
               #State_DwellAndReOx_SupplyToDeck:
                   IF #DECK_MANAGE_START_SUPPLY.ShutdownDemand THEN
                       #State.System := #State_Shutdown;
                   ELSIF "1092_HMI_OP_FLAGS".DeckSupplyOk THEN
                       #State.ReOx := #State_DwellAndReOx_OpenPVV;
                   ELSE
                       #DECK_MANAGE_START_SUPPLY();
                       "58_INTRNL_COMMS".BWT_TO_GCU.SPLY_GAS := True;
                       "58_INTRNL_COMMS".BWT_TO_GCU.STP_GAS := False;
                   END_IF;
               #State_DwellAndReOx_OpenPVV:
                   IF "1090_HMI_IP_FLAGS".PressVacuumValves THEN
                       #State.ReOx := #State_DwellAndReOx_OpenGTT;
                   ELSE
                       #NextStageCheck := "1151_NEXT_STAGE_CHECK_PVV"(AlarmState := #State_Shutdown, PVVX_OUT := #PVVX_OUT, State := #State, TankData := #TankData);
                       IF #NextStageCheck.Demand_Complete AND NOT #NextStageCheck.Alarm_Active THEN
                           #State.ReOx := #State_DwellAndReOx_OpenGTT;
                       END_IF;
                   END_IF;
               #State_DwellAndReOx_OpenGTT:
                   #NextStageCheck := "1150_NEXT_STAGE_CHECK_GTT"(AlarmState := #State_Shutdown, GTT_OUT := #GTT_OUT, State := #State, TankData := #TankData);
                   IF #NextStageCheck.Demand_Complete AND NOT #NextStageCheck.Alarm_Active THEN
                       #State.ReOx := #State_DwellAndReOx_Monitor;
                       "1134_MOVE_TANKS_INGROUP_NEW_STATE"(TankData := #TankData,
                                                          State := #State,
                                                          NewState := #TankState_ReOx);
                       // Reset timer information for this new treatment group
                       #XEOX_TIMER(IN := False,
                                   PT := "1190_FIXED_CONSTANTS".ReOxMin_Time,
                                   R := True);
                       #XEOX_PAUSE_TIMER(IN := False,
                                         PT := #MaxTimerPT,
                                         R := True);
                       #XEOX_PausedTime := LT#0s;
                   END_IF;
               #State_DwellAndReOx_Monitor:
                   IF #XEOX_TIMER.Q THEN
                       #NextStageCheck := "1153_NEXT_STAGE_CHECK_XEOX"(AlarmState := #State_Shutdown, State := #State, TankData := #TankData);
                       IF #NextStageCheck.Demand_Complete AND NOT #NextStageCheck.Alarm_Active THEN
                           #NextTreatmentGroup := "1136_CALC_NEXT_TREATMENT_GROUP"(NumberOfTreatmentGroups := "1190_FIXED_CONSTANTS".NumberOfTreatmentGroups, State := #State, TankData := #TankData);
                           IF #NextTreatmentGroup = -1 THEN
                               #DECK_MANAGE_STOP_SUPPLY.Stage := 0;
                               #State.ReOx := #State_DwellAndReOx_StopSupplyToDeck;
                           ELSE
                               #State.ReOx := #State_DwellAndReOx_CloseGTT;
                           END_IF;
                       END_IF;
                   ELSE
                       IF "58_INTRNL_COMMS".GCU_TO_BWT.GAS_AVLBL THEN
                           // continue counting on the reox timer as GCU is in a healthy state.
                           // increment the paused time as this shall be added to the deoxmin_time due to stoppage.
                           #XEOX_PausedTime += #XEOX_PAUSE_TIMER.ET;
                           #XEOX_TIMER(IN := True,
                                       PT := "1190_FIXED_CONSTANTS".ReOxMin_Time + #XEOX_PausedTime,
                                       R := False);
                           // keep XEOX pause timer in reset state.
                           #XEOX_PAUSE_TIMER(IN := False,
                                             PT := #MaxTimerPT,
                                             R := True);
                       ELSE
                           // Keep reox timer paused, whilst pause timer increments.
                           #XEOX_TIMER(IN := False,
                                       PT := "1190_FIXED_CONSTANTS".ReOxMin_Time + #XEOX_PausedTime,
                                       R := False);
                           #XEOX_PAUSE_TIMER(IN := True,
                                             PT := #MaxTimerPT,
                                             R := False);
                       END_IF;
                   END_IF;
               #State_DwellAndReOx_CloseGTT:
                   #NextStageCheck := "1150_NEXT_STAGE_CHECK_GTT"(AlarmState := #State_Shutdown, GTT_OUT := #GTT_OUT, State := #State, TankData := #TankData);
                   IF #NextStageCheck.Demand_Complete AND NOT #NextStageCheck.Alarm_Active THEN
                       // All tanks in this treatment group are now re-oxed, move them to post-dwell tank state.
                       "1134_MOVE_TANKS_INGROUP_NEW_STATE"(TankData := #TankData,
                                                          State := #State,
                                                          NewState := #TankState_PostDwell);
                      #NextTreatmentGroup := "1136_CALC_NEXT_TREATMENT_GROUP"(NumberOfTreatmentGroups := "1190_FIXED_CONSTANTS".NumberOfTreatmentGroups, State := #State, TankData := #TankData);
                       IF #NextTreatmentGroup = -1 THEN
                           #State.TreatmentGroup := 1;
                           #State.System := #State_DwellAndComplete;
                           #State.Complete := #State_DwellAndComplete_WaitPostDwell;
                       ELSE
                           // Are there more treatment groups to go? If so, restart the ReOx process on the next treatment group.
                           #State.TreatmentGroup := #NextTreatmentGroup;
                           #State.ReOx := #State_DwellAndReOx_WaitMidDwell;
                       END_IF;
                   END_IF;
               #State_DwellAndReOx_StopSupplyToDeck:
                   IF #DECK_MANAGE_STOP_SUPPLY.ShutdownDemand THEN
                       // Deck supply has failed, shutdown demand.
                       #State.System := #State_Shutdown;
                   ELSIF #DECK_MANAGE_STOP_SUPPLY.StopDeckSupplyDone THEN
                       // Deck stop supply is complete, go back to close the final set of GTT valves.
                       #State.ReOx := #State_DwellAndReOx_CloseGTT;
                   ELSE
                       // Deck stop supply is not complete yet, run stop supply to deck automation.
                       #DECK_MANAGE_STOP_SUPPLY();
                       "58_INTRNL_COMMS".BWT_TO_GCU.SPLY_GAS := False;
                       "58_INTRNL_COMMS".BWT_TO_GCU.STP_GAS := True;
                   END_IF;
           END_CASE;

       #State_DwellAndComplete:
           CASE #State.Complete OF
               #State_DwellAndComplete_WaitPostDwell:
                   #NextStageCheck := "1152_NEXT_STAGE_CHECK_TIMER"(AlarmState := #State_Shutdown, State := #State, TankData := #TankData);
                   IF #NextStageCheck.Demand_Complete AND NOT #NextStageCheck.Alarm_Active THEN
                       "1134_MOVE_TANKS_INGROUP_NEW_STATE"(TankData := #TankData,
                                                          State := #State,
                                                          NewState := #TankState_Done);
                      #NextTreatmentGroup := "1136_CALC_NEXT_TREATMENT_GROUP"(NumberOfTreatmentGroups := "1190_FIXED_CONSTANTS".NumberOfTreatmentGroups, State := #State, TankData := #TankData);
                       IF #NextTreatmentGroup = -1 THEN
                           #State.Complete := #State_DwellAndComplete_Done;
                       ELSE
                           // Are there more treatment groups to go? If so, wait for the next treatment group to finish post-dwell.
                           #State.TreatmentGroup := #NextTreatmentGroup;
                           #State.Complete := #State_DwellAndComplete_WaitPostDwell;
                       END_IF;
                   END_IF;
               #State_DwellAndComplete_Done:
                   // At this stage, all tanks have been processed.
                   "1092_HMI_OP_FLAGS".HMI_Warnings.Active := True;
                   "1092_HMI_OP_FLAGS".HMI_Warnings.Message := 'Ballast Water Treatment process has completed. All active tanks have been treated.';
           END_CASE;
       #State_Shutdown:
           "58_INTRNL_COMMS".BWT_TO_GCU.SHT_DN := True;
           IF #ShutdownStageReset THEN
               // If this is the first call to the shutdown, reset the stage to zero
               // do not call this reset again once called once.
               #DECK_MANAGE_STOP_SUPPLY.Stage := 0;
               #ShutdownStageReset := false;
           END_IF;
           IF #DECK_MANAGE_STOP_SUPPLY.ShutdownDemand THEN
               // Deck supply has failed, shutdown demand.6000
               #State.System := #State_Shutdown;
               "1092_HMI_OP_FLAGS".HMI_Warnings.Active := True;
               "1092_HMI_OP_FLAGS".HMI_Warnings.Message := 'BWTS Shutdown: failed to stop supply to main deck';
           ELSIF #DECK_MANAGE_STOP_SUPPLY.StopDeckSupplyDone THEN
               "1092_HMI_OP_FLAGS".HMI_Warnings.Active := True;
               "1092_HMI_OP_FLAGS".HMI_Warnings.Message := 'BWTS Shutdown: maain deck supply stopped';
           ELSE
               // Deck stop supply is not complete yet, run stop supply to deck automation.
               "1092_HMI_OP_FLAGS".HMI_Warnings.Active := True;
               "1092_HMI_OP_FLAGS".HMI_Warnings.Message := 'BWTS Shutdown: closing main line to deck';
               #DECK_MANAGE_STOP_SUPPLY();
           END_IF;
   END_CASE;

   (*
       Set all actuate commands to false to initialise on each scan cycle. Therefore each tank must now
       confirm that it wants the valve in question to actuate. Then call each tank in turn, make control
       decisions based on 1. The tank sub-state, the system operating state (and subsequently, deox/reox
       states if applicable.
   *)
   FOR #Index := 1 TO #NumberOfTanks DO
       #GTT_IN.GTT_Actuate[#Index] := False;
       #PVVX_IN.PVVx_Actuate[#Index] := False;
   END_FOR;
   #TANK_CONTROL_FPT(State := #State,
                     PVVX_IN := #PVVX_IN,
                     GTT_IN := #GTT_IN,
                     PVVX_OUT_DATA := #PVVX_OUT,
                     GTT_OUT_DATA := #GTT_OUT,
                     TankData := #TankData[1],
                     TankIPData := "20_TANKS_IP_DATA".RIO_01.FIRST_TANK);
   #TANK_CONTROL_1P(State := #State,
                    PVVX_IN := #PVVX_IN,
                    GTT_IN := #GTT_IN,
                    PVVX_OUT_DATA := #PVVX_OUT,
                    GTT_OUT_DATA := #GTT_OUT,
                    TankData := #TankData[2],
                    TankIPData := "20_TANKS_IP_DATA".RIO_01.SECOND_TANK);
   #TANK_CONTROL_1S(State := #State,
                    PVVX_IN := #PVVX_IN,
                    GTT_IN := #GTT_IN,
                    PVVX_OUT_DATA := #PVVX_OUT,
                    GTT_OUT_DATA := #GTT_OUT,
                    TankData := #TankData[3],
                    TankIPData := "20_TANKS_IP_DATA".RIO_01.THIRD_TANK);
   #TANK_CONTROL_2P(State := #State,
                    PVVX_IN := #PVVX_IN,
                    GTT_IN := #GTT_IN,
                    PVVX_OUT_DATA := #PVVX_OUT,
                    GTT_OUT_DATA := #GTT_OUT,
                    TankData := #TankData[4],
                    TankIPData := "20_TANKS_IP_DATA".RIO_02.FIRST_TANK);
   #TANK_CONTROL_2S(State := #State,
                    PVVX_IN := #PVVX_IN,
                    GTT_IN := #GTT_IN,
                    PVVX_OUT_DATA := #PVVX_OUT,
                    GTT_OUT_DATA := #GTT_OUT,
                    TankData := #TankData[5],
                    TankIPData := "20_TANKS_IP_DATA".RIO_02.SECOND_TANK);
   #TANK_CONTROL_3P(State := #State,
                    PVVX_IN := #PVVX_IN,
                    GTT_IN := #GTT_IN,
                    PVVX_OUT_DATA := #PVVX_OUT,
                    GTT_OUT_DATA := #GTT_OUT,
                    TankData := #TankData[6],
                    TankIPData := "20_TANKS_IP_DATA".RIO_03.FIRST_TANK);
   #TANK_CONTROL_3S(State := #State,
                    PVVX_IN := #PVVX_IN,
                    GTT_IN := #GTT_IN,
                    PVVX_OUT_DATA := #PVVX_OUT,
                    GTT_OUT_DATA := #GTT_OUT,
                    TankData := #TankData[7],
                    TankIPData := "20_TANKS_IP_DATA".RIO_03.SECOND_TANK);
   #TANK_CONTROL_4P(State := #State,
                    PVVX_IN := #PVVX_IN,
                    GTT_IN := #GTT_IN,
                    PVVX_OUT_DATA := #PVVX_OUT,
                    GTT_OUT_DATA := #GTT_OUT,
                    TankData := #TankData[8],
                    TankIPData := "20_TANKS_IP_DATA".RIO_04.FIRST_TANK);
   #TANK_CONTROL_4S(State := #State,
                    PVVX_IN := #PVVX_IN,
                    GTT_IN := #GTT_IN,
                    PVVX_OUT_DATA := #PVVX_OUT,
                    GTT_OUT_DATA := #GTT_OUT,
                    TankData := #TankData[9],
                    TankIPData := "20_TANKS_IP_DATA".RIO_04.SECOND_TANK);
   #TANK_CONTROL_5P(State := #State,
                    PVVX_IN := #PVVX_IN,
                    GTT_IN := #GTT_IN,
                    PVVX_OUT_DATA := #PVVX_OUT,
                    GTT_OUT_DATA := #GTT_OUT,
                    TankData := #TankData[10],
                    TankIPData := "20_TANKS_IP_DATA".RIO_05.FIRST_TANK);
   #TANK_CONTROL_5S(State := #State,
                    PVVX_IN := #PVVX_IN,
                    GTT_IN := #GTT_IN,
                    PVVX_OUT_DATA := #PVVX_OUT,
                    GTT_OUT_DATA := #GTT_OUT,
                    TankData := #TankData[11],
                    TankIPData := "20_TANKS_IP_DATA".RIO_05.SECOND_TANK);
   #TANK_CONTROL_6P(State := #State,
                    PVVX_IN := #PVVX_IN,
                    GTT_IN := #GTT_IN,
                    PVVX_OUT_DATA := #PVVX_OUT,
                    GTT_OUT_DATA := #GTT_OUT,
                    TankData := #TankData[12],
                    TankIPData := "20_TANKS_IP_DATA".RIO_06.FIRST_TANK);
   #TANK_CONTROL_6S(State := #State,
                    PVVX_IN := #PVVX_IN,
                    GTT_IN := #GTT_IN,
                    PVVX_OUT_DATA := #PVVX_OUT,
                    GTT_OUT_DATA := #GTT_OUT,
                    TankData := #TankData[13],
                    TankIPData := "20_TANKS_IP_DATA".RIO_06.SECOND_TANK);
   #TANK_CONTROL_APT(State := #State,
                     PVVX_IN := #PVVX_IN,
                     GTT_IN := #GTT_IN,
                     PVVX_OUT_DATA := #PVVX_OUT,
                     GTT_OUT_DATA := #GTT_OUT,
                     TankData := #TankData[14],
                     TankIPData := "20_TANKS_IP_DATA".RIO_07.FIRST_TANK);

   (*
       Management of the GTT valves and Vent valves (if applicable). Decisions on the valve management are made in
       the sub tank control, along with the main sequencer events. *_OUT data reports the demand completion status and alarms.
   *)
   #GTT_MANAGE_VALVES(GTT_Exclusivity := #GTT_Exclusivity,
                            GTT_IN := #GTT_IN,
                            GTT_OUT := #GTT_OUT);
   #PVV_MANAGE_VALVES(PVVX_IN := #PVVX_IN,
                      PVVX_OUT => #PVVX_OUT);

   // Push the state information to the GCU.
   "58_INTRNL_COMMS".BWT_TO_GCU.STATE := #State.System;
END_FUNCTION_BLOCK

FUNCTION_BLOCK "1101_RIO_MANUAL_CONTROL"   // FB1101, LAD
{ S7_Optimized_Access := 'TRUE' }
VERSION : 0.1
// Manual control maps HMI manual demand directly to the port controls for commisioning and testing purposes. This block is only run if the HMI has been set into Manual operating mode.
// 
// Feedback is produced through the normal channels in blocks 1110-1129.
BEGIN

REGION Network 1: RIO 01 (FPT) Manual valve control
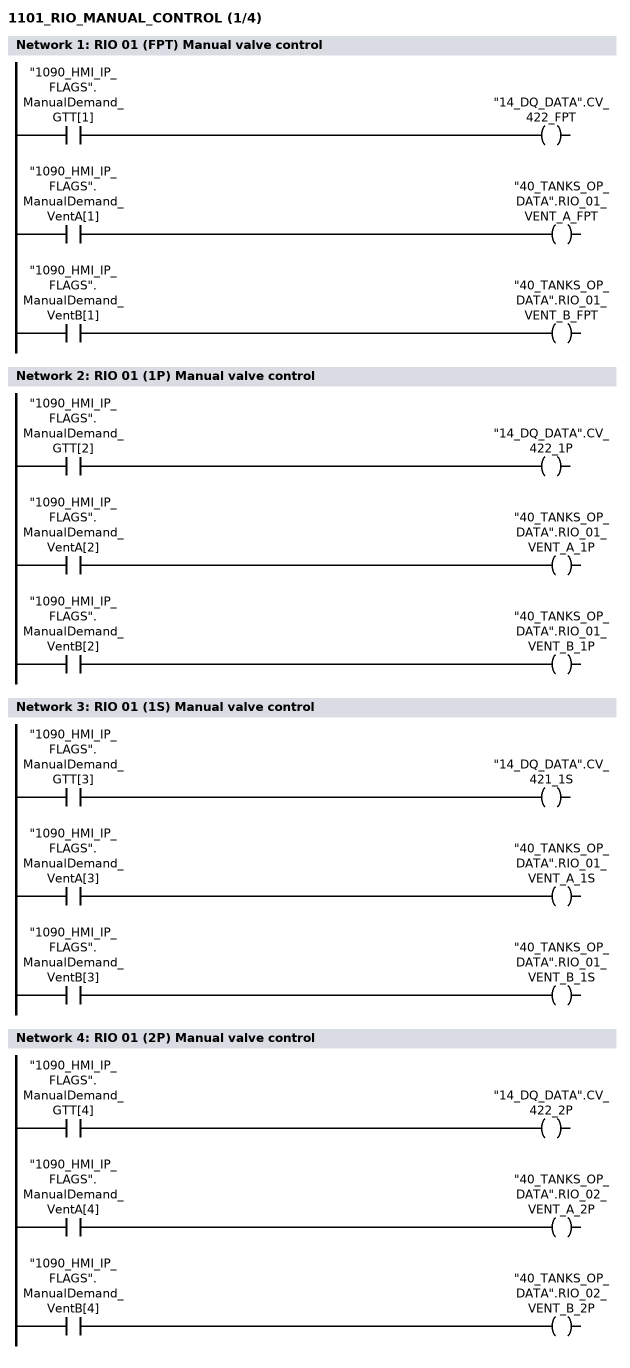
   RUNG wire#powerrail
      Contact( "1090_HMI_IP_FLAGS".ManualDemand_GTT[1] )
      Coil( "14_DQ_DATA".CV_422_FPT )
   END_RUNG
   RUNG wire#powerrail
      Contact( "1090_HMI_IP_FLAGS".ManualDemand_VentA[1] )
      Coil( "40_TANKS_OP_DATA".RIO_01_VENT_A_FPT )
   END_RUNG
   RUNG wire#powerrail
      Contact( "1090_HMI_IP_FLAGS".ManualDemand_VentB[1] )
      Coil( "40_TANKS_OP_DATA".RIO_01_VENT_B_FPT )
   END_RUNG
   // the same network as SCL:
   "14_DQ_DATA".CV_422_FPT := "1090_HMI_IP_FLAGS".ManualDemand_GTT[1];
   "40_TANKS_OP_DATA".RIO_01_VENT_A_FPT := "1090_HMI_IP_FLAGS".ManualDemand_VentA[1];
   "40_TANKS_OP_DATA".RIO_01_VENT_B_FPT := "1090_HMI_IP_FLAGS".ManualDemand_VentB[1];
END_REGION

REGION Network 2: RIO 01 (1P) Manual valve control
   RUNG wire#powerrail
      Contact( "1090_HMI_IP_FLAGS".ManualDemand_GTT[2] )
      Coil( "14_DQ_DATA".CV_422_1P )
   END_RUNG
   RUNG wire#powerrail
      Contact( "1090_HMI_IP_FLAGS".ManualDemand_VentA[2] )
      Coil( "40_TANKS_OP_DATA".RIO_01_VENT_A_1P )
   END_RUNG
   RUNG wire#powerrail
      Contact( "1090_HMI_IP_FLAGS".ManualDemand_VentB[2] )
      Coil( "40_TANKS_OP_DATA".RIO_01_VENT_B_1P )
   END_RUNG
   // the same network as SCL:
   "14_DQ_DATA".CV_422_1P := "1090_HMI_IP_FLAGS".ManualDemand_GTT[2];
   "40_TANKS_OP_DATA".RIO_01_VENT_A_1P := "1090_HMI_IP_FLAGS".ManualDemand_VentA[2];
   "40_TANKS_OP_DATA".RIO_01_VENT_B_1P := "1090_HMI_IP_FLAGS".ManualDemand_VentB[2];
END_REGION

REGION Network 3: RIO 01 (1S) Manual valve control
   RUNG wire#powerrail
      Contact( "1090_HMI_IP_FLAGS".ManualDemand_GTT[3] )
      Coil( "14_DQ_DATA".CV_421_1S )
   END_RUNG
   RUNG wire#powerrail
      Contact( "1090_HMI_IP_FLAGS".ManualDemand_VentA[3] )
      Coil( "40_TANKS_OP_DATA".RIO_01_VENT_A_1S )
   END_RUNG
   RUNG wire#powerrail
      Contact( "1090_HMI_IP_FLAGS".ManualDemand_VentB[3] )
      Coil( "40_TANKS_OP_DATA".RIO_01_VENT_B_1S )
   END_RUNG
   // the same network as SCL:
   "14_DQ_DATA".CV_421_1S := "1090_HMI_IP_FLAGS".ManualDemand_GTT[3];
   "40_TANKS_OP_DATA".RIO_01_VENT_A_1S := "1090_HMI_IP_FLAGS".ManualDemand_VentA[3];
   "40_TANKS_OP_DATA".RIO_01_VENT_B_1S := "1090_HMI_IP_FLAGS".ManualDemand_VentB[3];
END_REGION

REGION Network 4: RIO 01 (2P) Manual valve control
   RUNG wire#powerrail
      Contact( "1090_HMI_IP_FLAGS".ManualDemand_GTT[4] )
      Coil( "14_DQ_DATA".CV_422_2P )
   END_RUNG
   RUNG wire#powerrail
      Contact( "1090_HMI_IP_FLAGS".ManualDemand_VentA[4] )
      Coil( "40_TANKS_OP_DATA".RIO_02_VENT_A_2P )
   END_RUNG
   RUNG wire#powerrail
      Contact( "1090_HMI_IP_FLAGS".ManualDemand_VentB[4] )
      Coil( "40_TANKS_OP_DATA".RIO_02_VENT_B_2P )
   END_RUNG
   // the same network as SCL:
   "14_DQ_DATA".CV_422_2P := "1090_HMI_IP_FLAGS".ManualDemand_GTT[4];
   "40_TANKS_OP_DATA".RIO_02_VENT_A_2P := "1090_HMI_IP_FLAGS".ManualDemand_VentA[4];
   "40_TANKS_OP_DATA".RIO_02_VENT_B_2P := "1090_HMI_IP_FLAGS".ManualDemand_VentB[4];
END_REGION

REGION Network 5: RIO 01 (2S) Manual valve control
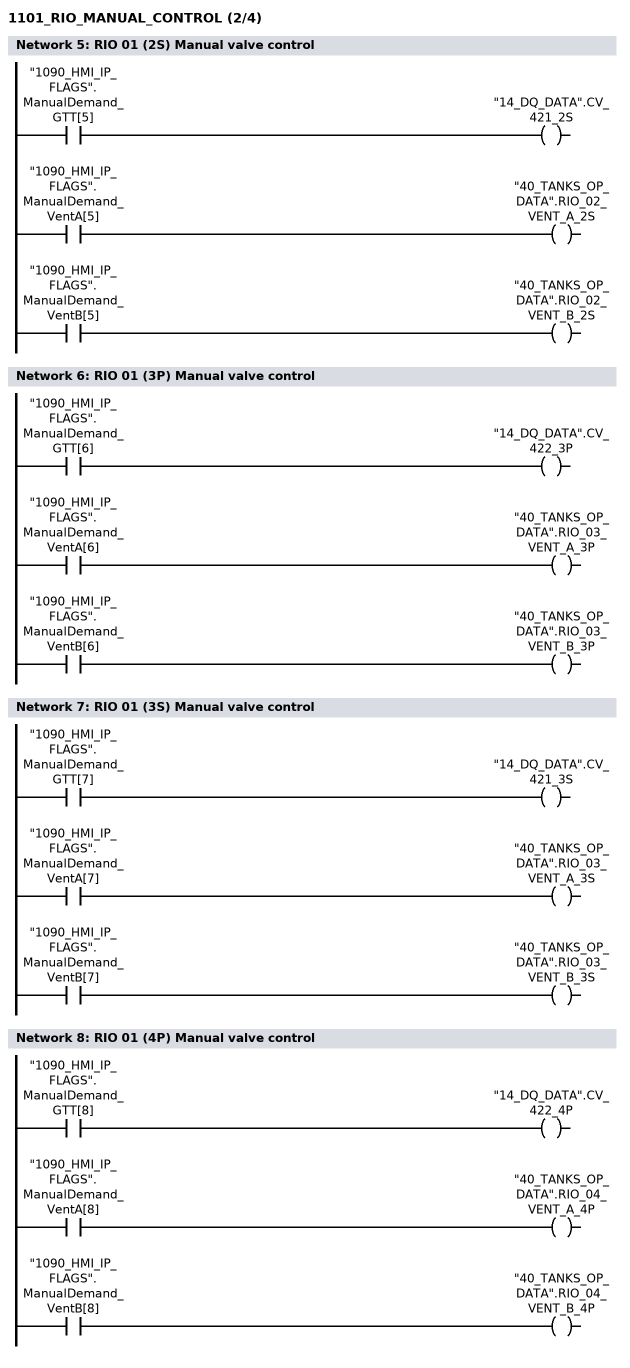
   RUNG wire#powerrail
      Contact( "1090_HMI_IP_FLAGS".ManualDemand_GTT[5] )
      Coil( "14_DQ_DATA".CV_421_2S )
   END_RUNG
   RUNG wire#powerrail
      Contact( "1090_HMI_IP_FLAGS".ManualDemand_VentA[5] )
      Coil( "40_TANKS_OP_DATA".RIO_02_VENT_A_2S )
   END_RUNG
   RUNG wire#powerrail
      Contact( "1090_HMI_IP_FLAGS".ManualDemand_VentB[5] )
      Coil( "40_TANKS_OP_DATA".RIO_02_VENT_B_2S )
   END_RUNG
   // the same network as SCL:
   "14_DQ_DATA".CV_421_2S := "1090_HMI_IP_FLAGS".ManualDemand_GTT[5];
   "40_TANKS_OP_DATA".RIO_02_VENT_A_2S := "1090_HMI_IP_FLAGS".ManualDemand_VentA[5];
   "40_TANKS_OP_DATA".RIO_02_VENT_B_2S := "1090_HMI_IP_FLAGS".ManualDemand_VentB[5];
END_REGION

REGION Network 6: RIO 01 (3P) Manual valve control
   RUNG wire#powerrail
      Contact( "1090_HMI_IP_FLAGS".ManualDemand_GTT[6] )
      Coil( "14_DQ_DATA".CV_422_3P )
   END_RUNG
   RUNG wire#powerrail
      Contact( "1090_HMI_IP_FLAGS".ManualDemand_VentA[6] )
      Coil( "40_TANKS_OP_DATA".RIO_03_VENT_A_3P )
   END_RUNG
   RUNG wire#powerrail
      Contact( "1090_HMI_IP_FLAGS".ManualDemand_VentB[6] )
      Coil( "40_TANKS_OP_DATA".RIO_03_VENT_B_3P )
   END_RUNG
   // the same network as SCL:
   "14_DQ_DATA".CV_422_3P := "1090_HMI_IP_FLAGS".ManualDemand_GTT[6];
   "40_TANKS_OP_DATA".RIO_03_VENT_A_3P := "1090_HMI_IP_FLAGS".ManualDemand_VentA[6];
   "40_TANKS_OP_DATA".RIO_03_VENT_B_3P := "1090_HMI_IP_FLAGS".ManualDemand_VentB[6];
END_REGION

REGION Network 7: RIO 01 (3S) Manual valve control
   RUNG wire#powerrail
      Contact( "1090_HMI_IP_FLAGS".ManualDemand_GTT[7] )
      Coil( "14_DQ_DATA".CV_421_3S )
   END_RUNG
   RUNG wire#powerrail
      Contact( "1090_HMI_IP_FLAGS".ManualDemand_VentA[7] )
      Coil( "40_TANKS_OP_DATA".RIO_03_VENT_A_3S )
   END_RUNG
   RUNG wire#powerrail
      Contact( "1090_HMI_IP_FLAGS".ManualDemand_VentB[7] )
      Coil( "40_TANKS_OP_DATA".RIO_03_VENT_B_3S )
   END_RUNG
   // the same network as SCL:
   "14_DQ_DATA".CV_421_3S := "1090_HMI_IP_FLAGS".ManualDemand_GTT[7];
   "40_TANKS_OP_DATA".RIO_03_VENT_A_3S := "1090_HMI_IP_FLAGS".ManualDemand_VentA[7];
   "40_TANKS_OP_DATA".RIO_03_VENT_B_3S := "1090_HMI_IP_FLAGS".ManualDemand_VentB[7];
END_REGION

REGION Network 8: RIO 01 (4P) Manual valve control
   RUNG wire#powerrail
      Contact( "1090_HMI_IP_FLAGS".ManualDemand_GTT[8] )
      Coil( "14_DQ_DATA".CV_422_4P )
   END_RUNG
   RUNG wire#powerrail
      Contact( "1090_HMI_IP_FLAGS".ManualDemand_VentA[8] )
      Coil( "40_TANKS_OP_DATA".RIO_04_VENT_A_4P )
   END_RUNG
   RUNG wire#powerrail
      Contact( "1090_HMI_IP_FLAGS".ManualDemand_VentB[8] )
      Coil( "40_TANKS_OP_DATA".RIO_04_VENT_B_4P )
   END_RUNG
   // the same network as SCL:
   "14_DQ_DATA".CV_422_4P := "1090_HMI_IP_FLAGS".ManualDemand_GTT[8];
   "40_TANKS_OP_DATA".RIO_04_VENT_A_4P := "1090_HMI_IP_FLAGS".ManualDemand_VentA[8];
   "40_TANKS_OP_DATA".RIO_04_VENT_B_4P := "1090_HMI_IP_FLAGS".ManualDemand_VentB[8];
END_REGION

REGION Network 9: RIO 01 (4S) Manual valve control
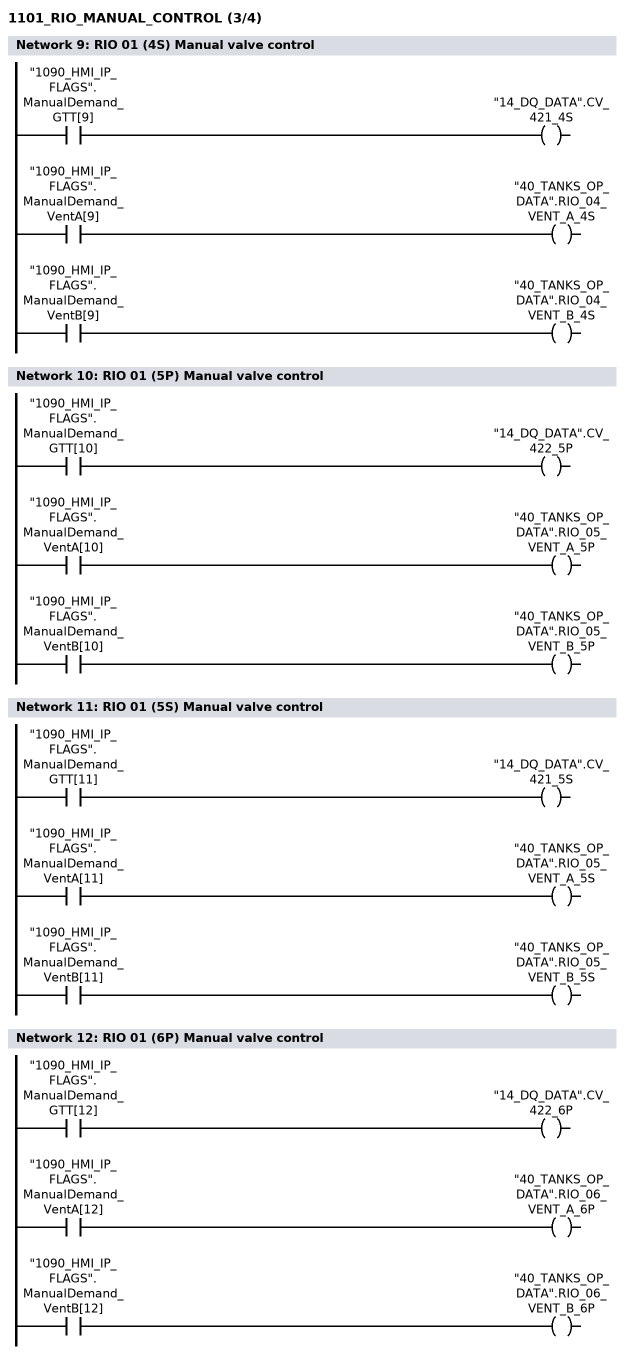
   RUNG wire#powerrail
      Contact( "1090_HMI_IP_FLAGS".ManualDemand_GTT[9] )
      Coil( "14_DQ_DATA".CV_421_4S )
   END_RUNG
   RUNG wire#powerrail
      Contact( "1090_HMI_IP_FLAGS".ManualDemand_VentA[9] )
      Coil( "40_TANKS_OP_DATA".RIO_04_VENT_A_4S )
   END_RUNG
   RUNG wire#powerrail
      Contact( "1090_HMI_IP_FLAGS".ManualDemand_VentB[9] )
      Coil( "40_TANKS_OP_DATA".RIO_04_VENT_B_4S )
   END_RUNG
   // the same network as SCL:
   "14_DQ_DATA".CV_421_4S := "1090_HMI_IP_FLAGS".ManualDemand_GTT[9];
   "40_TANKS_OP_DATA".RIO_04_VENT_A_4S := "1090_HMI_IP_FLAGS".ManualDemand_VentA[9];
   "40_TANKS_OP_DATA".RIO_04_VENT_B_4S := "1090_HMI_IP_FLAGS".ManualDemand_VentB[9];
END_REGION

REGION Network 10: RIO 01 (5P) Manual valve control
   RUNG wire#powerrail
      Contact( "1090_HMI_IP_FLAGS".ManualDemand_GTT[10] )
      Coil( "14_DQ_DATA".CV_422_5P )
   END_RUNG
   RUNG wire#powerrail
      Contact( "1090_HMI_IP_FLAGS".ManualDemand_VentA[10] )
      Coil( "40_TANKS_OP_DATA".RIO_05_VENT_A_5P )
   END_RUNG
   RUNG wire#powerrail
      Contact( "1090_HMI_IP_FLAGS".ManualDemand_VentB[10] )
      Coil( "40_TANKS_OP_DATA".RIO_05_VENT_B_5P )
   END_RUNG
   // the same network as SCL:
   "14_DQ_DATA".CV_422_5P := "1090_HMI_IP_FLAGS".ManualDemand_GTT[10];
   "40_TANKS_OP_DATA".RIO_05_VENT_A_5P := "1090_HMI_IP_FLAGS".ManualDemand_VentA[10];
   "40_TANKS_OP_DATA".RIO_05_VENT_B_5P := "1090_HMI_IP_FLAGS".ManualDemand_VentB[10];
END_REGION

REGION Network 11: RIO 01 (5S) Manual valve control
   RUNG wire#powerrail
      Contact( "1090_HMI_IP_FLAGS".ManualDemand_GTT[11] )
      Coil( "14_DQ_DATA".CV_421_5S )
   END_RUNG
   RUNG wire#powerrail
      Contact( "1090_HMI_IP_FLAGS".ManualDemand_VentA[11] )
      Coil( "40_TANKS_OP_DATA".RIO_05_VENT_A_5S )
   END_RUNG
   RUNG wire#powerrail
      Contact( "1090_HMI_IP_FLAGS".ManualDemand_VentB[11] )
      Coil( "40_TANKS_OP_DATA".RIO_05_VENT_B_5S )
   END_RUNG
   // the same network as SCL:
   "14_DQ_DATA".CV_421_5S := "1090_HMI_IP_FLAGS".ManualDemand_GTT[11];
   "40_TANKS_OP_DATA".RIO_05_VENT_A_5S := "1090_HMI_IP_FLAGS".ManualDemand_VentA[11];
   "40_TANKS_OP_DATA".RIO_05_VENT_B_5S := "1090_HMI_IP_FLAGS".ManualDemand_VentB[11];
END_REGION

REGION Network 12: RIO 01 (6P) Manual valve control
   RUNG wire#powerrail
      Contact( "1090_HMI_IP_FLAGS".ManualDemand_GTT[12] )
      Coil( "14_DQ_DATA".CV_422_6P )
   END_RUNG
   RUNG wire#powerrail
      Contact( "1090_HMI_IP_FLAGS".ManualDemand_VentA[12] )
      Coil( "40_TANKS_OP_DATA".RIO_06_VENT_A_6P )
   END_RUNG
   RUNG wire#powerrail
      Contact( "1090_HMI_IP_FLAGS".ManualDemand_VentB[12] )
      Coil( "40_TANKS_OP_DATA".RIO_06_VENT_B_6P )
   END_RUNG
   // the same network as SCL:
   "14_DQ_DATA".CV_422_6P := "1090_HMI_IP_FLAGS".ManualDemand_GTT[12];
   "40_TANKS_OP_DATA".RIO_06_VENT_A_6P := "1090_HMI_IP_FLAGS".ManualDemand_VentA[12];
   "40_TANKS_OP_DATA".RIO_06_VENT_B_6P := "1090_HMI_IP_FLAGS".ManualDemand_VentB[12];
END_REGION

REGION Network 13: RIO 01 (6S) Manual valve control
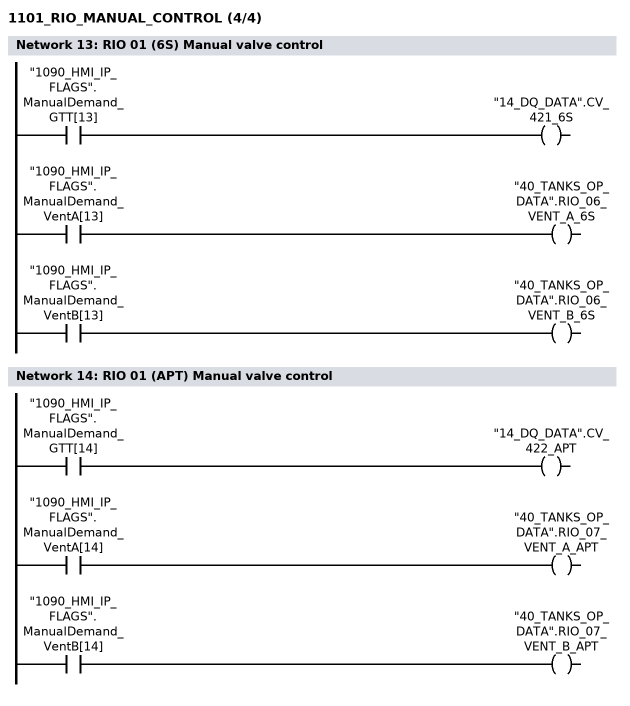
   RUNG wire#powerrail
      Contact( "1090_HMI_IP_FLAGS".ManualDemand_GTT[13] )
      Coil( "14_DQ_DATA".CV_421_6S )
   END_RUNG
   RUNG wire#powerrail
      Contact( "1090_HMI_IP_FLAGS".ManualDemand_VentA[13] )
      Coil( "40_TANKS_OP_DATA".RIO_06_VENT_A_6S )
   END_RUNG
   RUNG wire#powerrail
      Contact( "1090_HMI_IP_FLAGS".ManualDemand_VentB[13] )
      Coil( "40_TANKS_OP_DATA".RIO_06_VENT_B_6S )
   END_RUNG
   // the same network as SCL:
   "14_DQ_DATA".CV_421_6S := "1090_HMI_IP_FLAGS".ManualDemand_GTT[13];
   "40_TANKS_OP_DATA".RIO_06_VENT_A_6S := "1090_HMI_IP_FLAGS".ManualDemand_VentA[13];
   "40_TANKS_OP_DATA".RIO_06_VENT_B_6S := "1090_HMI_IP_FLAGS".ManualDemand_VentB[13];
END_REGION

REGION Network 14: RIO 01 (APT) Manual valve control
   RUNG wire#powerrail
      Contact( "1090_HMI_IP_FLAGS".ManualDemand_GTT[14] )
      Coil( "14_DQ_DATA".CV_422_APT )
   END_RUNG
   RUNG wire#powerrail
      Contact( "1090_HMI_IP_FLAGS".ManualDemand_VentA[14] )
      Coil( "40_TANKS_OP_DATA".RIO_07_VENT_A_APT )
   END_RUNG
   RUNG wire#powerrail
      Contact( "1090_HMI_IP_FLAGS".ManualDemand_VentB[14] )
      Coil( "40_TANKS_OP_DATA".RIO_07_VENT_B_APT )
   END_RUNG
   // the same network as SCL:
   "14_DQ_DATA".CV_422_APT := "1090_HMI_IP_FLAGS".ManualDemand_GTT[14];
   "40_TANKS_OP_DATA".RIO_07_VENT_A_APT := "1090_HMI_IP_FLAGS".ManualDemand_VentA[14];
   "40_TANKS_OP_DATA".RIO_07_VENT_B_APT := "1090_HMI_IP_FLAGS".ManualDemand_VentB[14];
END_REGION
END_FUNCTION_BLOCK

// folder: 1000 - 1999 BWT System Control/1105 - 1109 Main Control

FUNCTION_BLOCK "1105_TANK_CONTROL"   // FB1105, SCL
{ S7_Optimized_Access := 'TRUE' }
VERSION : 0.1
   VAR_INPUT
      State : "SYSTEM_STATES";   // State information on this tank instantiated.
      TankIPData : "TANK_IP_DATA";   // Tank input data from the RIO/Tank associated with this instantiated tank.
      PVVX_OUT_DATA : "VALVE_PVVX_OUT";
      GTT_OUT_DATA : "VALVE_GTT_OUT";
   END_VAR
   VAR_IN_OUT
      TankData : "TANK_DATA";   // Combined tank data for the tank which this instantiated object refers to.
      PVVX_IN : "VALVE_PVVX_IN";
      GTT_IN : "VALVE_GTT_IN";
   END_VAR
   VAR RETAIN
      DWELL_TIMER : TONR_LTIME;   // Timer for measuring Mid-Dwell or Post-Dwell process. Combined to reduce complexity of next stage checking. Processes are split by states so are mutually exclusive.
      MONITOR_TIMER : TONR_LTIME;
      ReOx_InitialTargetpHLevelAchieved : Bool;
   END_VAR
   VAR CONSTANT
      State_Init : Int := 0;   // State for initialization
      State_PreDwell : Int := 1;   // State to control pre-dwell
      State_DeOx : Int := 2;   // State to control DeOx and mid-dwell
      State_DeOx_SupplyToDeck : Int := 200;
      State_DeOx_ClosePVV : Int := 201;
      State_DeOx_OpenGTT : Int := 202;
      State_DeOx_Monitor : Int := 203;
      State_DeOx_CloseGTT : Int := 204;
      State_DeOx_StopSupplyToDeck : Int := 205;
      State_DwellAndReOx : Int := 3;   // State to control ReOx and post-dwell
      State_DwellAndReOx_WaitMidDwell : Int := 300;
      State_DwellAndReOx_SupplyToDeck : Int := 301;
      State_DwellAndReOx_OpenPVV : Int := 302;
      State_DwellAndReOx_OpenGTT : Int := 303;
      State_DwellAndReOx_Monitor : Int := 304;
      State_DwellAndReOx_CloseGTT : Int := 305;
      State_DwellAndReOx_StopSupplyToDeck : Int := 306;
      State_DwellAndComplete : Int := 4;
      State_DwellAndComplete_WaitPostDwell : Int := 400;
      State_DwellAndComplete_Done : Int := 401;
      State_Shutdown : Int := 5;   // State to control shutdown events
      TankState_Init : Int := 1000;
      TankState_PreDwell : Int := 1001;
      TankState_DeOx : Int := 1002;
      TankState_MidDwell : Int := 1003;
      TankState_ReOx : Int := 1004;
      TankState_PostDwell : Int := 1005;
      TankState_Done : Int := 1006;
   END_VAR
BEGIN
   // NOTE: TANK_CONTROL cannot modify its own state, but can report it has completed its current operation.
   // Only the top level sequencer may modify the state of a sub-tank.

